// TIA Portal project "Urban Intersection Control System" (V17)

(* hardware
DEVICE "S7-1500/ET200MP station_1"  S7-1500 station
   slot 0: "Rail_0"  Rack  6ES7 590-1***0-0AA0
   slot 1: "PLC_UICS_01"  CPU 1512C-1 PN  6ES7 512-1CK00-0AB0  V2.9
      slot 3: "CPU display_1"  6ES7591-1AA00-0AA0
      slot 32768: "PROFINET interface_1"  X1
         slot 32769: "Port_1"  X1 P1
         slot 32770: "Port_2"  X1 P2
      slot 34817: "Virtual CP interface port_1"  Virtual CP interface port  Virtual CP interface port
DEVICE "HMI_1"  KTP1200 Basic PN
   slot 0: "HMI_1"  KTP1200 Basic PN  6AV2 123-2MB03-0AX0  17.0.0.0
   slot 1: "HMI_RT_1"  KTP1200 Basic PN  6AV2 123-2MB03-0AX0  17.0.0.0
   slot 5: "HMI_1.IE_CP_1"  PROFINET Interface  17.0.0.0
      slot 1: "PROFINET Interface_1"  PROFINET Interface
         slot 1: "Port_1"  Port
*)

// ===== PLC "PLC_UICS_01"  CPU 1512C-1 PN =====

VAR_GLOBAL   // PLC tag table "UICS_Table"
   "PB_Ped_Main" AT %I10.2 : Bool;   // Push button for pedestrian crossing on Main Street
   "PB_Ped_Cross" AT %I10.3 : Bool;   // Push button for pedestrian crossing on Cross Street
   "EM_Main_Override" AT %I10.4 : Bool;   // Emergency override signal (e.g. ambulances) on Main Street
   "EM_Cross_Override" AT %I10.5 : Bool;   // Emergency override signal on Cross Street
   "SENSOR_Main_Vehicle" AT %I10.6 : Bool;   // Vehicle detection sensor on Main Street
   "SENSOR_Cross_Vehicle" AT %I10.7 : Bool;   // Vehicle detection sensor on Cross Street
   "TL_Main_Red_West" AT %Q4.0 : Bool;   // Red traffic light signal for western Main Street
   "TL_Main_Yellow_West" AT %Q4.2 : Bool;   // Yellow traffic light signal for western Main Street
   "TL_Main_Green_West" AT %Q4.4 : Bool;   // Green traffic light signal for western Main Street
   "TL_Cross_Red_North" AT %Q4.6 : Bool;   // Red traffic light signal for northern Cross Street
   "TL_Cross_Yellow_North" AT %Q5.0 : Bool;   // Yellow traffic light signal for northern Cross Street
   "TL_Cross_Green_North" AT %Q5.2 : Bool;   // Green traffic light signal for northern Cross Street
   "PED_Main_Walk_West" AT %Q5.4 : Bool;   // Pedestrian walk signal for western Main Street
   "PED_Main_DontWalk_West" AT %Q5.6 : Bool;   // Pedestrian don’t-walk signal for western Main Street
   "PED_Cross_Walk_North" AT %Q6.0 : Bool;   // Pedestrian walk signal for northern Cross Street
   "PED_Cross_DontWalk_North" AT %Q6.2 : Bool;   // Pedestrian don’t-walk signal for northern Cross Street
   "PED_Warning_Buzzer" AT %Q6.4 : Bool;   // Audible alert for pedestrian crossing
   "SYS_Stop" AT %I10.1 : Bool;   // Emergency stop function
   "SYS_Start" AT %I10.0 : Bool;   // Begins the system
   "TL_Main_Red_East" AT %Q4.1 : Bool;   // Red traffic light signal for eastern Main Street
   "TL_Main_Yellow_East" AT %Q4.3 : Bool;   // Yellow traffic light signal for eastern Main Street
   "TL_Main_Green_East" AT %Q4.5 : Bool;   // Green traffic light signal for eastern Main Street
   "TL_Cross_Red_South" AT %Q4.7 : Bool;   // Red traffic light signal for southern Cross Street
   "TL_Cross_Yellow_South" AT %Q5.1 : Bool;   // Yellow traffic light signal for southern Cross Street
   "TL_Cross_Green_South" AT %Q5.3 : Bool;   // Green traffic light signal for southern Cross Street
   "PED_Main_Walk_East" AT %Q5.5 : Bool;   // Pedestrian walk signal for eastern Main Street
   "PED_Main_DontWalk_East" AT %Q5.7 : Bool;   // Pedestrian don’t-walk signal for eastern Main Street
   "PED_Cross_Walk_South" AT %Q6.1 : Bool;   // Pedestrian walk signal for southern Cross Street
   "PED_Cross_DontWalk_South" AT %Q6.3 : Bool;   // Pedestrian don’t-walk signal for southern Cross Street
END_VAR

DATA_BLOCK "Main_Control_System_DB"   // DB1
{ S7_Optimized_Access := 'TRUE' }
VERSION : 0.1
// stored: InstanceOfName Main_Control_System
"Main_Control_System"
BEGIN
END_DATA_BLOCK

DATA_BLOCK "Traffic_Light_Operations_DB"   // DB3
{ S7_Optimized_Access := 'TRUE' }
VERSION : 0.1
// stored: InstanceOfName Traffic_Light_Operations
"Traffic_Light_Operations"
BEGIN
END_DATA_BLOCK

DATA_BLOCK "Status_Reset_DB"   // DB7
{ S7_Optimized_Access := 'TRUE' }
VERSION : 0.1
// stored: InstanceOfName Status_Reset
"Status_Reset"
BEGIN
END_DATA_BLOCK

// folder: System blocks/Program resources

DATA_BLOCK "Eastern_MainSt_Timer_DB"   // DB2
{ S7_Optimized_Access := 'TRUE' }
AUTHOR : Simatic
FAMILY : IEC
NAME : IEC_TMR
VERSION : 1.0
// stored: InstanceOfName IEC_TIMER
"IEC_TIMER"
BEGIN
END_DATA_BLOCK

DATA_BLOCK "Western_MainSt_Timer_DB"   // DB4
{ S7_Optimized_Access := 'TRUE' }
AUTHOR : Simatic
FAMILY : IEC
NAME : IEC_TMR
VERSION : 1.0
// stored: InstanceOfName IEC_TIMER
"IEC_TIMER"
BEGIN
END_DATA_BLOCK

DATA_BLOCK "Southern_CrossSt_Timer_DB"   // DB5
{ S7_Optimized_Access := 'TRUE' }
AUTHOR : Simatic
FAMILY : IEC
NAME : IEC_TMR
VERSION : 1.0
// stored: InstanceOfName IEC_TIMER
"IEC_TIMER"
BEGIN
END_DATA_BLOCK

DATA_BLOCK "Northern_CrossSt_Timer_DB"   // DB6
{ S7_Optimized_Access := 'TRUE' }
AUTHOR : Simatic
FAMILY : IEC
NAME : IEC_TMR
VERSION : 1.0
// stored: InstanceOfName IEC_TIMER
"IEC_TIMER"
BEGIN
END_DATA_BLOCK

// folder: (top level)

FUNCTION_BLOCK "Main_Control_System"   // FB1, LAD
{ S7_Optimized_Access := 'TRUE' }
VERSION : 0.1
   VAR_INPUT
      System_Start : Bool;   // Activates the system
      System_Stop : Bool;   // Emergency stop function
   END_VAR
   VAR
      System_Latch : Bool;   // Allows the system to remain active after initially starting up
      System_Running : Bool;   // System is actively running
      Emergency_Stop : Bool;   // Emergency stop activated flag
      HMI_Start_Command : Bool;   // Allows HMI to start the system
      HMI_Stop_Command : Bool;   // Allows HMI to stop the system
      HMI_Latch_Command : Bool;   // Allows HMI visualization to remain active after initially starting up
      HMI_Run_Command : Bool;   // Allows HMI to run the system
   END_VAR
BEGIN

REGION Network 1: System Start
   // Starts the system if all conditions are met
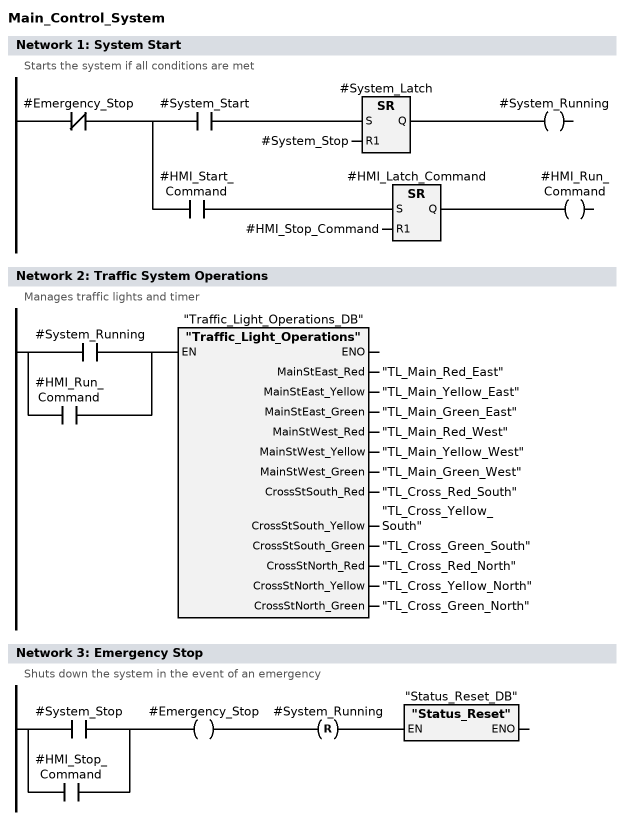
   RUNG wire#powerrail
      I_Contact( #Emergency_Stop )
      wire#w1
      Contact( #System_Start )
      S_SR(operand := #System_Latch, r1 := #System_Stop)
      Coil( #System_Running )
   END_RUNG
   RUNG wire#w1
      Contact( #HMI_Start_Command )
      S_SR(operand := #HMI_Latch_Command, r1 := #HMI_Stop_Command)
      Coil( #HMI_Run_Command )
   END_RUNG
   // the same network as SCL:
   IF NOT #Emergency_Stop AND #System_Start THEN
       #System_Latch := TRUE;   // SR flip-flop
   END_IF;
   IF #System_Stop THEN #System_Latch := FALSE; END_IF;
   #System_Running := #System_Latch;
   IF NOT #Emergency_Stop AND #HMI_Start_Command THEN
       #HMI_Latch_Command := TRUE;   // SR flip-flop
   END_IF;
   IF #HMI_Stop_Command THEN #HMI_Latch_Command := FALSE; END_IF;
   #HMI_Run_Command := #HMI_Latch_Command;
END_REGION

REGION Network 2: Traffic System Operations
   // Manages traffic lights and timer
   RUNG wire#powerrail
      Contact( #System_Running )
      wire#w1
      "Traffic_Light_Operations_DB"(MainStEast_Red => "TL_Main_Red_East", MainStEast_Yellow => "TL_Main_Yellow_East", MainStEast_Green => "TL_Main_Green_East", MainStWest_Red => "TL_Main_Red_West", MainStWest_Yellow => "TL_Main_Yellow_West", MainStWest_Green => "TL_Main_Green_West", CrossStSouth_Red => "TL_Cross_Red_South", CrossStSouth_Yellow => "TL_Cross_Yellow_South", CrossStSouth_Green => "TL_Cross_Green_South", CrossStNorth_Red => "TL_Cross_Red_North", CrossStNorth_Yellow => "TL_Cross_Yellow_North", CrossStNorth_Green => "TL_Cross_Green_North")
   END_RUNG
   RUNG wire#powerrail
      Contact( #HMI_Run_Command )
   END_RUNG wire#w1
   // the same network as SCL:
   IF #System_Running OR #HMI_Run_Command THEN
       "Traffic_Light_Operations_DB"(MainStEast_Red => "TL_Main_Red_East",   // "Traffic_Light_Operations"
                               MainStEast_Yellow => "TL_Main_Yellow_East",
                               MainStEast_Green => "TL_Main_Green_East",
                               MainStWest_Red => "TL_Main_Red_West",
                               MainStWest_Yellow => "TL_Main_Yellow_West",
                               MainStWest_Green => "TL_Main_Green_West",
                               CrossStSouth_Red => "TL_Cross_Red_South",
                               CrossStSouth_Yellow => "TL_Cross_Yellow_South",
                               CrossStSouth_Green => "TL_Cross_Green_South",
                               CrossStNorth_Red => "TL_Cross_Red_North",
                               CrossStNorth_Yellow => "TL_Cross_Yellow_North",
                               CrossStNorth_Green => "TL_Cross_Green_North");
   END_IF;
END_REGION

REGION Network 3: Emergency Stop
   // Shuts down the system in the event of an emergency
   RUNG wire#powerrail
      Contact( #System_Stop )
      wire#w1
      Coil( #Emergency_Stop )
      R_Coil( #System_Running )
      "Status_Reset_DB"()
   END_RUNG
   RUNG wire#powerrail
      Contact( #HMI_Stop_Command )
   END_RUNG wire#w1
   // the same network as SCL:
   #Emergency_Stop := #System_Stop OR #HMI_Stop_Command;
   IF #Emergency_Stop THEN
       #System_Running := FALSE;
       "Status_Reset_DB"();   // "Status_Reset"
   END_IF;
END_REGION
END_FUNCTION_BLOCK

FUNCTION_BLOCK "Traffic_Light_Operations"   // FB2, LAD
{ S7_Optimized_Access := 'TRUE' }
VERSION : 0.1
   VAR_OUTPUT
      MainStEast_Red : Bool;   // Red traffic light signal for eastern Main Street
      MainStEast_Yellow : Bool;   // Yellow traffic light signal for eastern Main Street
      MainStEast_Green : Bool;   // Green traffic light signal for eastern Main Street
      MainStWest_Red : Bool;   // Red traffic light signal for western Main Street
      MainStWest_Yellow : Bool;   // Yellow traffic light signal for western Main Street
      MainStWest_Green : Bool;   // Green traffic light signal for western Main Street
      CrossStSouth_Red : Bool;   // Red traffic light signal for southern Cross Street
      CrossStSouth_Yellow : Bool;   // Yellow traffic light signal for southern Cross Street
      CrossStSouth_Green : Bool;   // Green traffic light signal for southern Cross Street
      CrossStNorth_Red : Bool;   // Red traffic light signal for northern Cross Street
      CrossStNorth_Yellow : Bool;   // Yellow traffic light signal for northern Cross Street
      CrossStNorth_Green : Bool;   // Green traffic light signal for northern Cross Street
   END_VAR
   VAR
      Traffic_Operations_Step : Int;   // Controls the state of traffic operations
      Eastern_MainSt_Seconds : Int;   // Allows HMI to read eastern Main Street traffic time
      Western_MainSt_Seconds : Int;   // Allows HMI to read western Main Street traffic time
      Southern_CrossSt_Seconds : Int;   // Allows HMI to read southern Cross Street traffic time
      Northern_CrossSt_Seconds : Int;   // Allows HMI to read northern Cross Street traffic time
      Initialize_Operation : Bool;   // Initiates traffic operations
   END_VAR
   VAR_TEMP
      Eastern_MainSt_ET_DInt : DInt;
      Eastern_MainSt_ET_Div : DInt;
      Western_MainSt_ET_DInt : DInt;
      Western_MainSt_ET_Div : DInt;
      Southern_CrossSt_ET_DInt : DInt;
      Southern_CrossSt_ET_Div : DInt;
      Northern_CrossSt_ET_DInt : DInt;
      Northern_CrossSt_ET_Div : DInt;
   END_VAR
   VAR_TEMP   // added for the SCL form of the ladder/FBD networks
      _w1 : Bool;
   END_VAR
BEGIN

REGION Network 1: Red Light Control
   // Organization of red traffic lights for Main Street and Cross Street
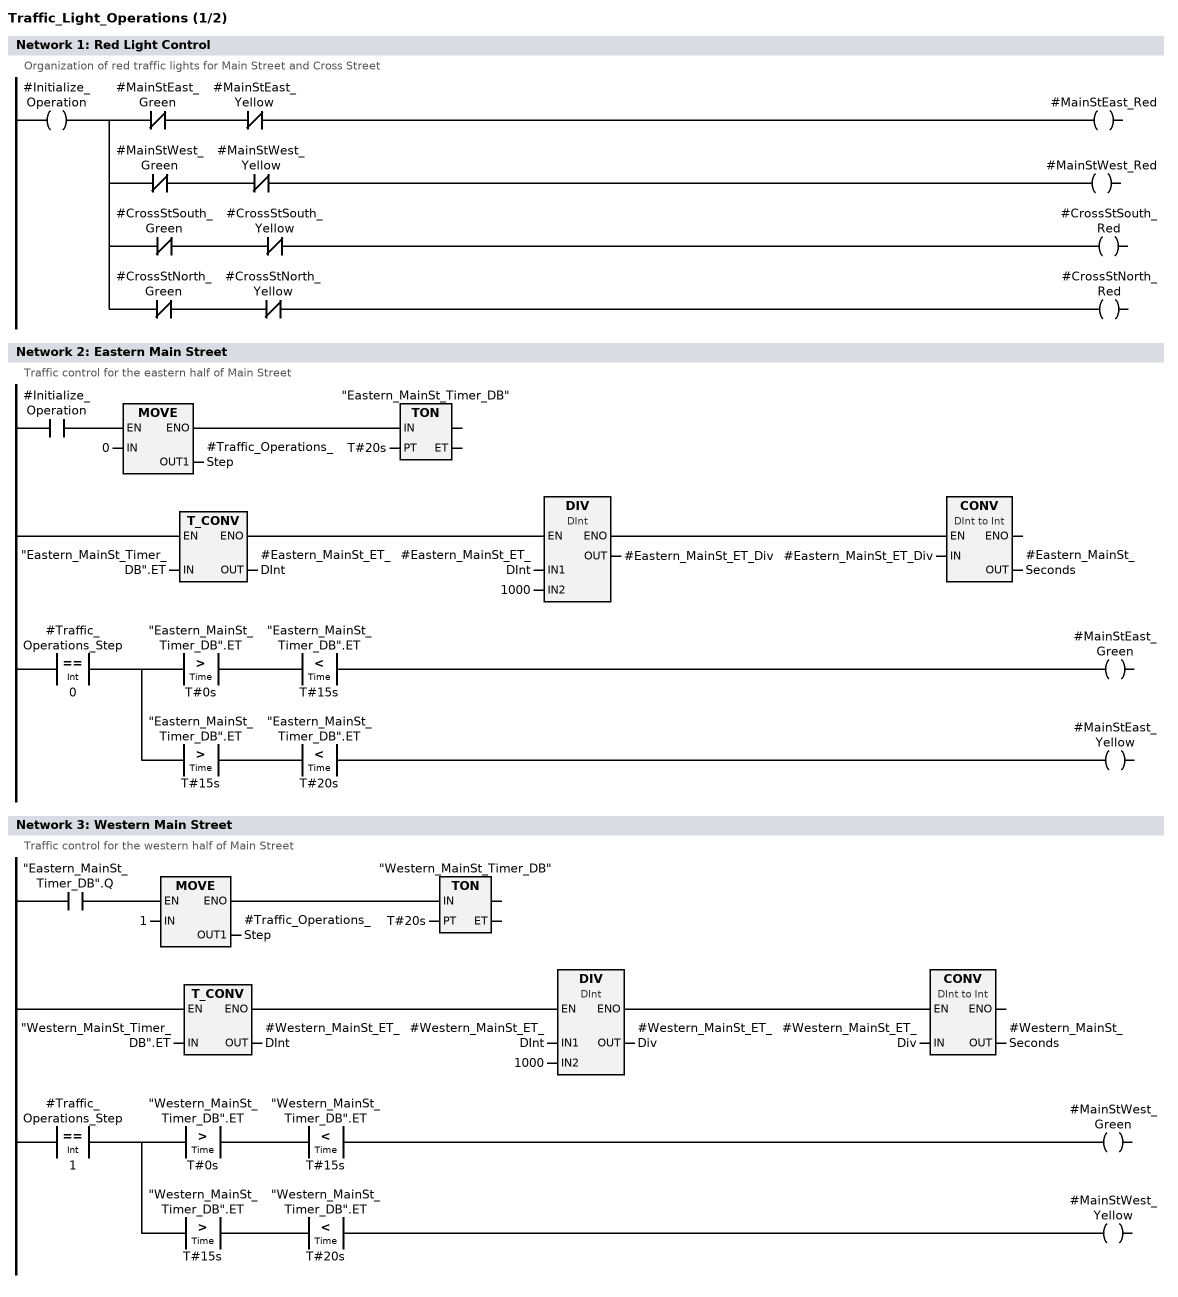
   RUNG wire#powerrail
      Coil( #Initialize_Operation )
      wire#w1
      I_Contact( #MainStEast_Green )
      I_Contact( #MainStEast_Yellow )
      Coil( #MainStEast_Red )
   END_RUNG
   RUNG wire#w1
      I_Contact( #MainStWest_Green )
      I_Contact( #MainStWest_Yellow )
      Coil( #MainStWest_Red )
   END_RUNG
   RUNG wire#w1
      I_Contact( #CrossStSouth_Green )
      I_Contact( #CrossStSouth_Yellow )
      Coil( #CrossStSouth_Red )
   END_RUNG
   RUNG wire#w1
      I_Contact( #CrossStNorth_Green )
      I_Contact( #CrossStNorth_Yellow )
      Coil( #CrossStNorth_Red )
   END_RUNG
   // the same network as SCL:
   #Initialize_Operation := TRUE;
   #MainStEast_Red := NOT #MainStEast_Green AND NOT #MainStEast_Yellow;
   #MainStWest_Red := NOT #MainStWest_Green AND NOT #MainStWest_Yellow;
   #CrossStSouth_Red := NOT #CrossStSouth_Green AND NOT #CrossStSouth_Yellow;
   #CrossStNorth_Red := NOT #CrossStNorth_Green AND NOT #CrossStNorth_Yellow;
END_REGION

REGION Network 2: Eastern Main Street
   // Traffic control for the eastern half of Main Street
   // ENO of a box is taken as its EN; it also drops when the box reports an error
   IF #Initialize_Operation THEN #Traffic_Operations_Step := 0; END_IF;
   "Eastern_MainSt_Timer_DB".TON(IN := #Initialize_Operation, PT := T#20s);
   #Eastern_MainSt_ET_DInt := T_CONV(IN := "Eastern_MainSt_Timer_DB".ET);
   #Eastern_MainSt_ET_Div := #Eastern_MainSt_ET_DInt / 1000;
   #Eastern_MainSt_Seconds := DINT_TO_INT(#Eastern_MainSt_ET_Div);
   #_w1 := #Traffic_Operations_Step = 0;
   #MainStEast_Green := #_w1 AND ("Eastern_MainSt_Timer_DB".ET > T#0s) AND ("Eastern_MainSt_Timer_DB".ET < T#15s);
   #MainStEast_Yellow := #_w1 AND ("Eastern_MainSt_Timer_DB".ET > T#15s) AND ("Eastern_MainSt_Timer_DB".ET < T#20s);
END_REGION

REGION Network 3: Western Main Street
   // Traffic control for the western half of Main Street
   // ENO of a box is taken as its EN; it also drops when the box reports an error
   IF "Eastern_MainSt_Timer_DB".Q THEN #Traffic_Operations_Step := 1; END_IF;
   "Western_MainSt_Timer_DB".TON(IN := "Eastern_MainSt_Timer_DB".Q, PT := T#20s);
   #Western_MainSt_ET_DInt := T_CONV(IN := "Western_MainSt_Timer_DB".ET);
   #Western_MainSt_ET_Div := #Western_MainSt_ET_DInt / 1000;
   #Western_MainSt_Seconds := DINT_TO_INT(#Western_MainSt_ET_Div);
   #_w1 := #Traffic_Operations_Step = 1;
   #MainStWest_Green := #_w1 AND ("Western_MainSt_Timer_DB".ET > T#0s) AND ("Western_MainSt_Timer_DB".ET < T#15s);
   #MainStWest_Yellow := #_w1 AND ("Western_MainSt_Timer_DB".ET > T#15s) AND ("Western_MainSt_Timer_DB".ET < T#20s);
END_REGION

REGION Network 4: Southern Cross Street
   // Traffic control for the southern half of Cross Street
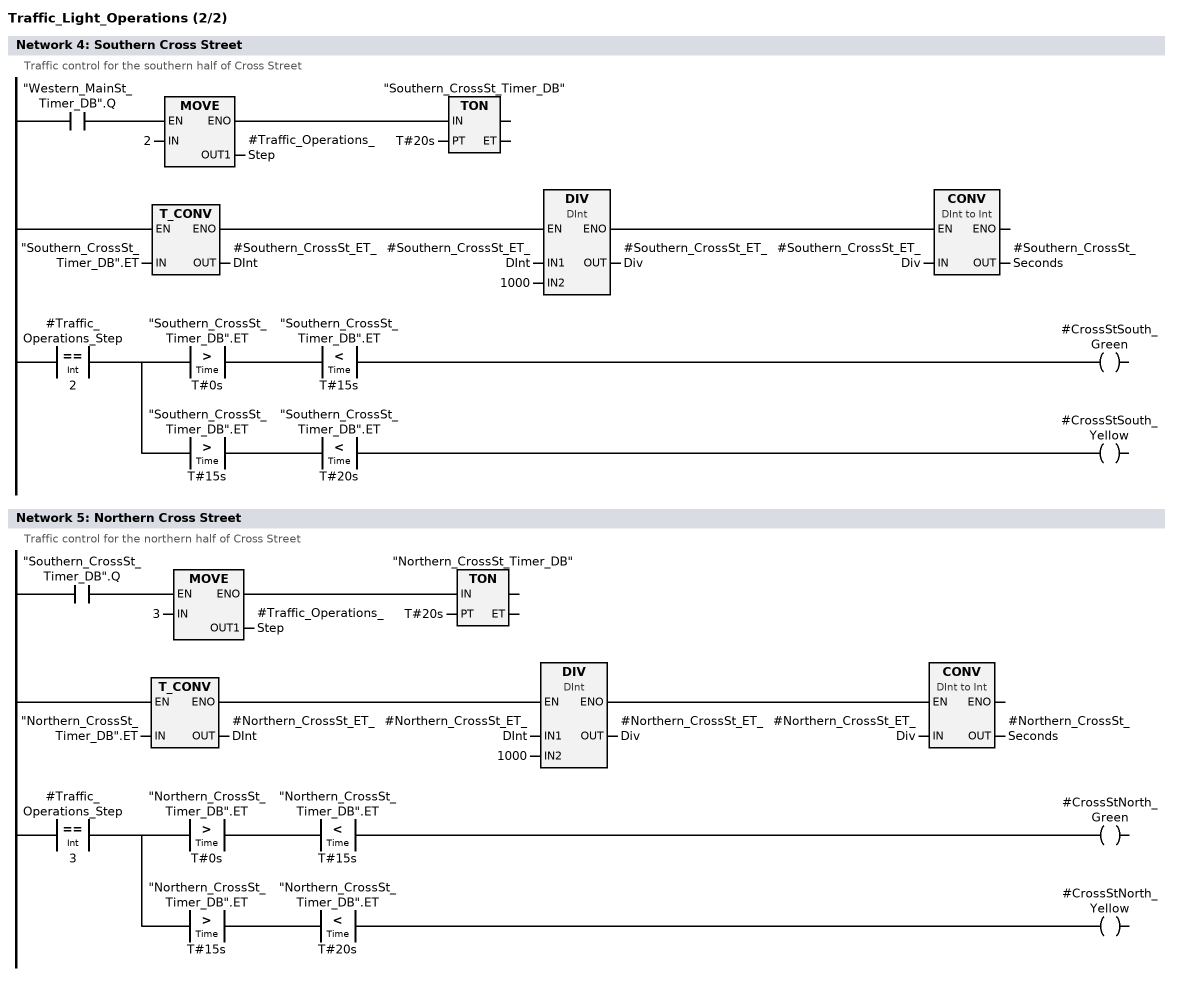
   // ENO of a box is taken as its EN; it also drops when the box reports an error
   IF "Western_MainSt_Timer_DB".Q THEN #Traffic_Operations_Step := 2; END_IF;
   "Southern_CrossSt_Timer_DB".TON(IN := "Western_MainSt_Timer_DB".Q, PT := T#20s);
   #Southern_CrossSt_ET_DInt := T_CONV(IN := "Southern_CrossSt_Timer_DB".ET);
   #Southern_CrossSt_ET_Div := #Southern_CrossSt_ET_DInt / 1000;
   #Southern_CrossSt_Seconds := DINT_TO_INT(#Southern_CrossSt_ET_Div);
   #_w1 := #Traffic_Operations_Step = 2;
   #CrossStSouth_Green := #_w1 AND ("Southern_CrossSt_Timer_DB".ET > T#0s) AND ("Southern_CrossSt_Timer_DB".ET < T#15s);
   #CrossStSouth_Yellow := #_w1 AND ("Southern_CrossSt_Timer_DB".ET > T#15s) AND ("Southern_CrossSt_Timer_DB".ET < T#20s);
END_REGION

REGION Network 5: Northern Cross Street
   // Traffic control for the northern half of Cross Street
   // ENO of a box is taken as its EN; it also drops when the box reports an error
   IF "Southern_CrossSt_Timer_DB".Q THEN #Traffic_Operations_Step := 3; END_IF;
   "Northern_CrossSt_Timer_DB".TON(IN := "Southern_CrossSt_Timer_DB".Q, PT := T#20s);
   #Northern_CrossSt_ET_DInt := T_CONV(IN := "Northern_CrossSt_Timer_DB".ET);
   #Northern_CrossSt_ET_Div := #Northern_CrossSt_ET_DInt / 1000;
   #Northern_CrossSt_Seconds := DINT_TO_INT(#Northern_CrossSt_ET_Div);
   #_w1 := #Traffic_Operations_Step = 3;
   #CrossStNorth_Green := #_w1 AND ("Northern_CrossSt_Timer_DB".ET > T#0s) AND ("Northern_CrossSt_Timer_DB".ET < T#15s);
   #CrossStNorth_Yellow := #_w1 AND ("Northern_CrossSt_Timer_DB".ET > T#15s) AND ("Northern_CrossSt_Timer_DB".ET < T#20s);
END_REGION
END_FUNCTION_BLOCK

FUNCTION_BLOCK "Status_Reset"   // FB3, LAD
{ S7_Optimized_Access := 'TRUE' }
VERSION : 0.1
BEGIN

REGION Network 1
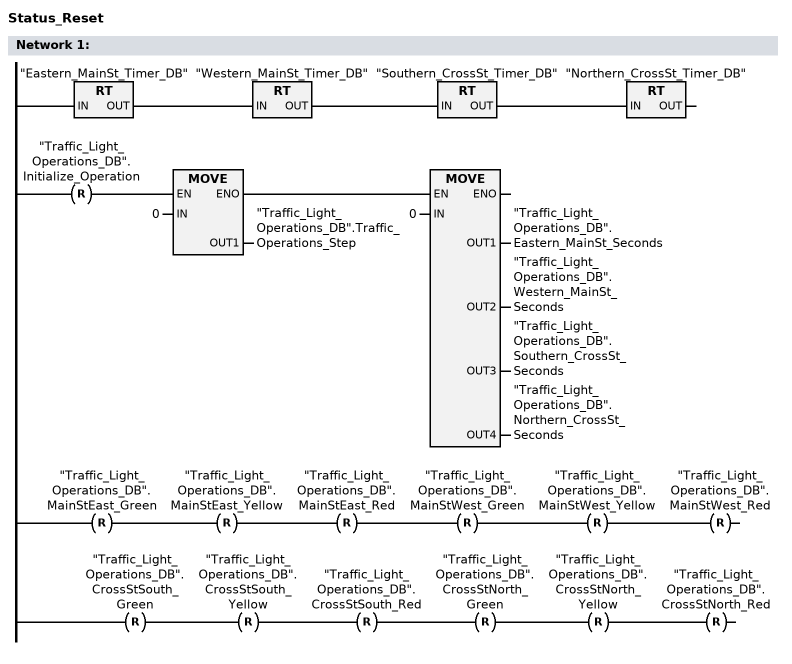
   RUNG wire#powerrail
      RT_Coil( "Eastern_MainSt_Timer_DB" )
      RT_Coil( "Western_MainSt_Timer_DB" )
      RT_Coil( "Southern_CrossSt_Timer_DB" )
      RT_Coil( "Northern_CrossSt_Timer_DB" )
   END_RUNG
   RUNG wire#powerrail
      R_Coil( "Traffic_Light_Operations_DB".Initialize_Operation )
      Move(in := 0, out1 => "Traffic_Light_Operations_DB".Traffic_Operations_Step)
      Move(in := 0, out1 => "Traffic_Light_Operations_DB".Eastern_MainSt_Seconds, out2 => "Traffic_Light_Operations_DB".Western_MainSt_Seconds, out3 => "Traffic_Light_Operations_DB".Southern_CrossSt_Seconds, out4 => "Traffic_Light_Operations_DB".Northern_CrossSt_Seconds)
   END_RUNG
   RUNG wire#powerrail
      R_Coil( "Traffic_Light_Operations_DB".MainStEast_Green )
      R_Coil( "Traffic_Light_Operations_DB".MainStEast_Yellow )
      R_Coil( "Traffic_Light_Operations_DB".MainStEast_Red )
      R_Coil( "Traffic_Light_Operations_DB".MainStWest_Green )
      R_Coil( "Traffic_Light_Operations_DB".MainStWest_Yellow )
      R_Coil( "Traffic_Light_Operations_DB".MainStWest_Red )
   END_RUNG
   RUNG wire#powerrail
      R_Coil( "Traffic_Light_Operations_DB".CrossStSouth_Green )
      R_Coil( "Traffic_Light_Operations_DB".CrossStSouth_Yellow )
      R_Coil( "Traffic_Light_Operations_DB".CrossStSouth_Red )
      R_Coil( "Traffic_Light_Operations_DB".CrossStNorth_Green )
      R_Coil( "Traffic_Light_Operations_DB".CrossStNorth_Yellow )
      R_Coil( "Traffic_Light_Operations_DB".CrossStNorth_Red )
   END_RUNG
   // the same network as SCL:
   RESET_TIMER("Eastern_MainSt_Timer_DB");
   RESET_TIMER("Western_MainSt_Timer_DB");
   RESET_TIMER("Southern_CrossSt_Timer_DB");
   RESET_TIMER("Northern_CrossSt_Timer_DB");
   "Traffic_Light_Operations_DB".Initialize_Operation := FALSE;
   "Traffic_Light_Operations_DB".Traffic_Operations_Step := 0;
   "Traffic_Light_Operations_DB".Eastern_MainSt_Seconds := 0;
   "Traffic_Light_Operations_DB".Western_MainSt_Seconds := 0;
   "Traffic_Light_Operations_DB".Southern_CrossSt_Seconds := 0;
   "Traffic_Light_Operations_DB".Northern_CrossSt_Seconds := 0;
   "Traffic_Light_Operations_DB".MainStEast_Green := FALSE;
   "Traffic_Light_Operations_DB".MainStEast_Yellow := FALSE;
   "Traffic_Light_Operations_DB".MainStEast_Red := FALSE;
   "Traffic_Light_Operations_DB".MainStWest_Green := FALSE;
   "Traffic_Light_Operations_DB".MainStWest_Yellow := FALSE;
   "Traffic_Light_Operations_DB".MainStWest_Red := FALSE;
   "Traffic_Light_Operations_DB".CrossStSouth_Green := FALSE;
   "Traffic_Light_Operations_DB".CrossStSouth_Yellow := FALSE;
   "Traffic_Light_Operations_DB".CrossStSouth_Red := FALSE;
   "Traffic_Light_Operations_DB".CrossStNorth_Green := FALSE;
   "Traffic_Light_Operations_DB".CrossStNorth_Yellow := FALSE;
   "Traffic_Light_Operations_DB".CrossStNorth_Red := FALSE;
END_REGION
END_FUNCTION_BLOCK

ORGANIZATION_BLOCK "Main"   // OB1, LAD, ProgramCycle
TITLE = "Main Program Sweep (Cycle)"
{ S7_Optimized_Access := 'TRUE' }
VERSION : 0.1
   VAR_INPUT
      Initial_Call : Bool;   // Initial call of this OB
      Remanence : Bool;   // =True, if remanent data are available
   END_VAR
BEGIN

REGION Network 1: Main
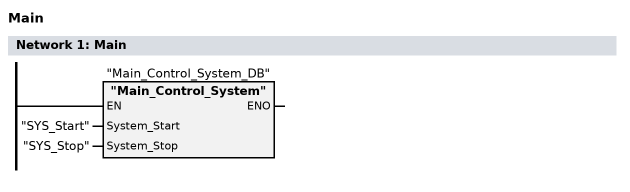
   RUNG wire#powerrail
      "Main_Control_System_DB"(System_Start := "SYS_Start", System_Stop := "SYS_Stop")
   END_RUNG
   // the same network as SCL:
   "Main_Control_System_DB"(System_Start := "SYS_Start", System_Stop := "SYS_Stop");   // "Main_Control_System"
END_REGION
END_ORGANIZATION_BLOCK

(* ===== HMI "HMI_RT_1" =====
system functions are stored by id; their names below are inferred from use
connection "HMI_Connection": ETHERNET, SMART_S7_1500_OMS

HMI tags "Default tag table"
   "Tag_ScreenNumber" : UInt, internal

HMI tags "UICS_HMI_Table"
   "MainStEast_RedLight" : Bool = PLC Traffic_Light_Operations_DB.MainStEast_Red AT %DB1.DBX0.0, 100 ms
   "MainStEast_YellowLight" : Bool = PLC Traffic_Light_Operations_DB.MainStEast_Yellow AT %DB1.DBX0.0, 100 ms
   "MainStEast_GreenLight" : Bool = PLC Traffic_Light_Operations_DB.MainStEast_Green AT %DB1.DBX0.0, 100 ms
   "MainStWest_RedLight" : Bool = PLC Traffic_Light_Operations_DB.MainStWest_Red AT %DB1.DBX0.0, 100 ms
   "MainStWest_YellowLight" : Bool = PLC Traffic_Light_Operations_DB.MainStWest_Yellow AT %DB1.DBX0.0, 100 ms
   "MainStWest_GreenLight" : Bool = PLC Traffic_Light_Operations_DB.MainStWest_Green AT %DB1.DBX0.0, 100 ms
   "CrossStSouth_RedLight" : Bool = PLC Traffic_Light_Operations_DB.CrossStSouth_Red AT %DB1.DBX0.0, 100 ms
   "CrossStSouth_YellowLight" : Bool = PLC Traffic_Light_Operations_DB.CrossStSouth_Yellow AT %DB1.DBX0.0, 100 ms
   "CrossStSouth_GreenLight" : Bool = PLC Traffic_Light_Operations_DB.CrossStSouth_Green AT %DB1.DBX0.0, 100 ms
   "CrossStNorth_RedLight" : Bool = PLC Traffic_Light_Operations_DB.CrossStNorth_Red AT %DB1.DBX0.0, 100 ms
   "CrossStNorth_YellowLight" : Bool = PLC Traffic_Light_Operations_DB.CrossStNorth_Yellow AT %DB1.DBX0.0, 100 ms
   "CrossStNorth_GreenLight" : Bool = PLC Traffic_Light_Operations_DB.CrossStNorth_Green AT %DB1.DBX0.0, 100 ms
   "Eastern_MainSt_Seconds" : Int = PLC Traffic_Light_Operations_DB.Eastern_MainSt_Seconds AT %DB1.DBX0.0, 100 ms
   "System_Running" : Bool = PLC Main_Control_System_DB.HMI_Run_Command AT %DB1.DBW0, 100 ms
   "Emergency_Stop" : Bool = PLC Main_Control_System_DB.Emergency_Stop AT %DB1.DBW0, 100 ms
   "Push_Button_Start" : Bool = PLC Main_Control_System_DB.HMI_Start_Command AT %DB1.DBX0.0, 100 ms
   "Push_Button_Stop" : Bool = PLC Main_Control_System_DB.HMI_Stop_Command AT %DB1.DBX0.0, 100 ms
   "Western_MainSt_Seconds" : Int = PLC Traffic_Light_Operations_DB.Western_MainSt_Seconds AT %DB1.DBW0, 100 ms
   "Southern_CrossSt_Seconds" : Int = PLC Traffic_Light_Operations_DB.Southern_CrossSt_Seconds AT %DB1.DBW0, 100 ms
   "Northern_CrossSt_Seconds" : Int = PLC Traffic_Light_Operations_DB.Northern_CrossSt_Seconds AT %DB1.DBW0, 100 ms

Template "Template_1" 1280x800
   Button "Exit" at 1182,752 size 67x47; TextOff 'Exit'; PictureOff "ExitRuntime_KTP1200_Basic_PN_TR"; PictureOn "ExitRuntime_KTP1200_Basic_PN_TR"
      on Release: StopRuntime(0)
   Button "Template_Button" at 1054,752 size 67x47; TextOff 'Text'
   Button "Template_Button_1" at 926,752 size 67x47; TextOff 'Text'
   Button "Template_Button_2" at 798,752 size 67x47; TextOff 'Text'
   Button "Template_Button_3" at 670,752 size 67x47; TextOff 'Text'
   Button "Template_Button_4" at 542,752 size 67x47; TextOff 'Text'
   Button "Template_Button_5" at 414,752 size 67x47; TextOff 'Text'
   Button "Template_Button_6" at 286,752 size 67x47; TextOff 'Text'
   Button "Alarms" at 158,752 size 67x47; TextOff 'Alarms'; PictureOff "AlarmDisplay_KTP1200_Basic_PN_TR"; PictureOn "AlarmDisplay_KTP1200_Basic_PN_TR"
      on Release: function_ef3f5d25("Alarm window_Unacknowledged", -1)
   Button "Start screen" at 30,752 size 67x47; TextOff 'Start screen'; PictureOff "NavigateHome_KTP1200_Basic_PN_TR"; PictureOn "NavigateHome_KTP1200_Basic_PN_TR"
      on Release: ActivateScreen("Root screen", 0)
   SymbolicIOField "Symbolic_IO_Field_Screen" at 87,9 size 1086x30; TextOff '0'; TextOn '1'; TextList "TextList_ScreenNames"
      ProcessValue <- "Tag_ScreenNumber"
      on Change: ActivateScreenByNumber("Tag_ScreenNumber", 0)
   DateTimeField "HmiScreenItemData" at 1175,24 size 105x24
   DateTimeField "HmiScreenItemData_1" at 1175,0 size 105x24
   GraphicView "Logo" at 0,0 size 85x48; Picture "Logo of HMI_1"

screen "Root screen" 1280x800, template "Template_1"
   on GenerateScreen: SetTag("Tag_ScreenNumber", 1)
   TextField "HmiScreenItemData" at 128,384 size 1024x27; Text 'Welcome to HMI_1 (KTP1200 Basic+ PN)!'

screen "Screen_1" 1280x800
   GraphicView "Four_Way_Road" at 319,94 size 612x612; Picture "Graphic_2"
   Group "MainStWest_TL" at 455,398 size 50x100
   Group "CrossStSouth_TL" at 622,509 size 100x50
   Group "CrossStNorth_TL" at 524,224 size 100x50
   IOField "I/O field_1" at 1057,314 size 96x32; FormatPattern s99; Unit  s
      ProcessValue <- "Eastern_MainSt_Seconds"
   Button "Button_1" at 25,569 size 96x32; TextOff 'Start'
      on Press: InvertBit("Push_Button_Start")
   Button "Button_2" at 190,569 size 96x32; TextOff 'Stop'
      on Press: InvertBit("Push_Button_Stop")
   Switch "Pushbutton_Square_G" at 47,619 size 50x50; CaptionText 'Switch'; TextOff '0'; TextOn '1'; PictureOff "Pushbutton_Square_G_Off_256c"; PictureOn "Pushbutton_Square_G_On_256c"
      ProcessValue <- "System_Running"
   Switch "Pushbutton_Square_R" at 211,619 size 50x50; CaptionText 'Switch'; TextOff '0'; TextOn '1'; PictureOff "Pushbutton_Square_R_Off_256c"; PictureOn "Pushbutton_Square_R_On_256c"
      ProcessValue <- "Emergency_Stop"
   Group "MainStEast_TL" at 751,301 size 50x100
   IOField "I/O field_2" at 576,50 size 96x32; FormatPattern s99; Unit  s
      ProcessValue <- "Northern_CrossSt_Seconds"
   IOField "I/O field_3" at 100,377 size 96x32; FormatPattern s99; Unit  s
      ProcessValue <- "Western_MainSt_Seconds"
   IOField "I/O field_4" at 577,752 size 96x32; FormatPattern s99; Unit  s
      ProcessValue <- "Southern_CrossSt_Seconds"
   TextField "Text field_1" at 505,22 size 263x25; Text 'Northern Cross St Traffic Time'
   TextField "Text field_2" at 33,345 size 263x25; Text 'Western Main St Traffic Time'
   TextField "Text field_5" at 987,281 size 263x25; Text 'Eastern Main St Traffic Time'
   TextField "Text field_6" at 516,724 size 263x25; Text 'Southern Cross St Traffic Time'
   Circle "Green_East" at 763,370 size 26x26
      Appearance <- "MainStEast_GreenLight"
   Circle "Red_East" at 763,310 size 26x26
      Appearance <- "MainStEast_RedLight"
   Circle "Yellow_East" at 763,340 size 26x26
      Appearance <- "MainStEast_YellowLight"
   Circle "Red_West" at 467,407 size 26x26
      Appearance <- "MainStWest_RedLight"
   Circle "Yellow_West" at 467,437 size 26x26
      Appearance <- "MainStWest_YellowLight"
   Circle "Green_West" at 467,467 size 26x26
      Appearance <- "MainStWest_GreenLight"
   Circle "Red_South" at 687,521 size 26x26
      Appearance <- "CrossStSouth_RedLight"
   Circle "Yellow_South" at 657,521 size 26x26
      Appearance <- "CrossStSouth_YellowLight"
   Circle "Green_South" at 627,521 size 26x26
      Appearance <- "CrossStSouth_GreenLight"
   Circle "Red_North" at 589,236 size 26x26
      Appearance <- "CrossStNorth_RedLight"
   Circle "Yellow_North" at 559,236 size 26x26
      Appearance <- "CrossStNorth_YellowLight"
   Circle "Green_North" at 529,236 size 26x26
      Appearance <- "CrossStNorth_GreenLight"
*)